
REGION Network 27: State 20 = Failed Ignition Attempt
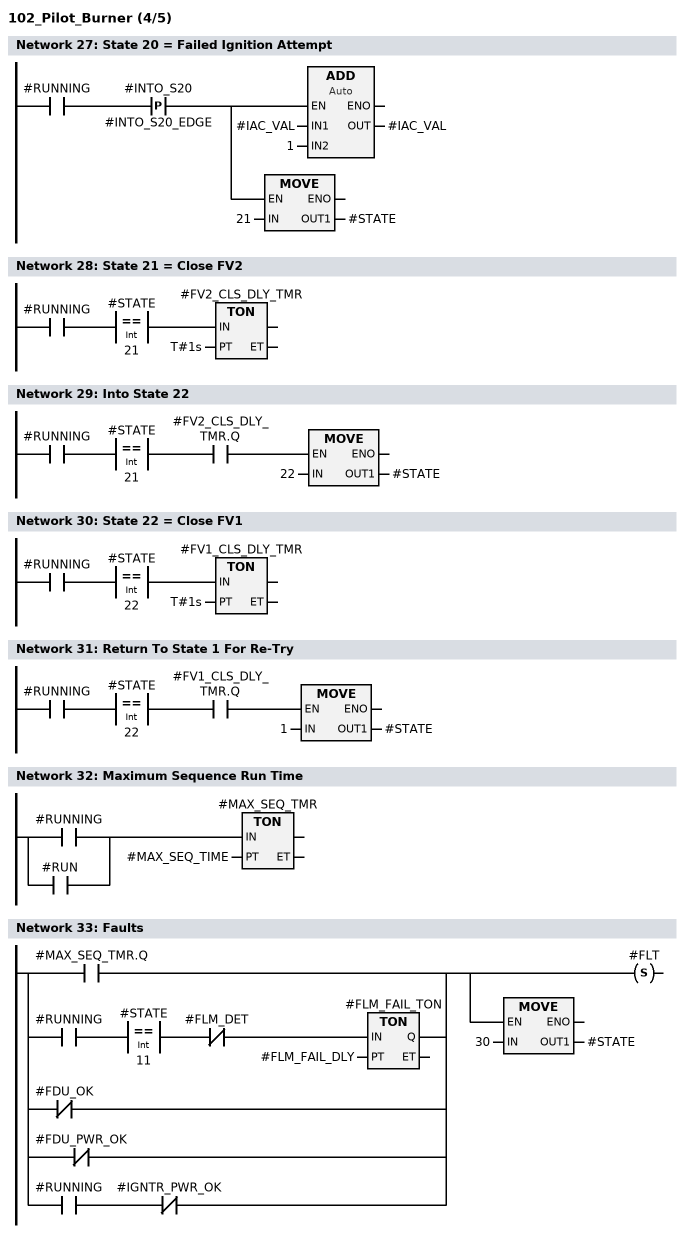
   RUNG wire#powerrail
      Contact( #RUNNING )
      P_Contact(operand := #INTO_S20, bit := #INTO_S20_EDGE)
      wire#w1
      Add(in1 := #IAC_VAL, in2 := 1, out => #IAC_VAL)
   END_RUNG
   RUNG wire#w1
      Move(in := 21, out1 => #STATE)
   END_RUNG
   // the same network as SCL:
   #_w1 := #RUNNING AND #INTO_S20 AND NOT #INTO_S20_EDGE;   // rising edge of #INTO_S20
   #INTO_S20_EDGE := #INTO_S20;
   IF #_w1 THEN
       #IAC_VAL := #IAC_VAL + 1;
       #STATE := 21;
   END_IF;
END_REGION

REGION Network 28: State 21 = Close FV2
   #FV2_CLS_DLY_TMR(IN := #RUNNING AND (#STATE = 21), PT := T#1s);   // TON
END_REGION

REGION Network 29: Into State 22
   RUNG wire#powerrail
      Contact( #RUNNING )
      { S7_Templates := "SrcType := Int" } EQ_Contact(in1 := #STATE, in2 := 21)
      Contact( #FV2_CLS_DLY_TMR.Q )
      Move(in := 22, out1 => #STATE)
   END_RUNG
   // the same network as SCL:
   IF #RUNNING AND (#STATE = 21) AND #FV2_CLS_DLY_TMR.Q THEN #STATE := 22; END_IF;
END_REGION

REGION Network 30: State 22 = Close FV1
   #FV1_CLS_DLY_TMR(IN := #RUNNING AND (#STATE = 22), PT := T#1s);   // TON
END_REGION

REGION Network 31: Return To State 1 For Re-Try
   RUNG wire#powerrail
      Contact( #RUNNING )
      { S7_Templates := "SrcType := Int" } EQ_Contact(in1 := #STATE, in2 := 22)
      Contact( #FV1_CLS_DLY_TMR.Q )
      Move(in := 1, out1 => #STATE)
   END_RUNG
   // the same network as SCL:
   IF #RUNNING AND (#STATE = 22) AND #FV1_CLS_DLY_TMR.Q THEN #STATE := 1; END_IF;
END_REGION

REGION Network 32: Maximum Sequence Run Time
   #MAX_SEQ_TMR(IN := #RUNNING OR #RUN, PT := #MAX_SEQ_TIME);   // TON
END_REGION

REGION Network 33: Faults
   #FLM_FAIL_TON(IN := #RUNNING AND (#STATE = 11) AND NOT #FLM_DET, PT := #FLM_FAIL_DLY);   // TON
   IF #MAX_SEQ_TMR.Q OR #FLM_FAIL_TON.Q OR NOT #FDU_OK OR NOT #FDU_PWR_OK OR (#RUNNING AND NOT #IGNTR_PWR_OK) THEN
       #FLT := TRUE;
       #STATE := 30;
   END_IF;
END_REGION

REGION Network 34: Reset Flag
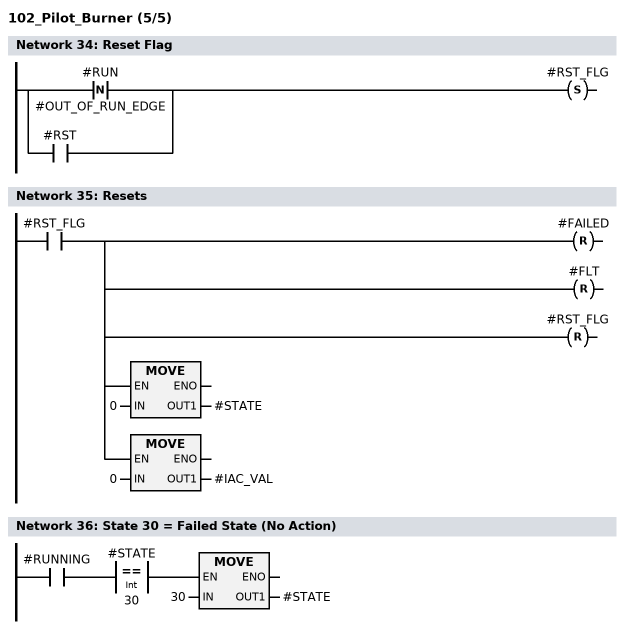
   RUNG wire#powerrail
      N_Contact(operand := #RUN, bit := #OUT_OF_RUN_EDGE)
      wire#w1
      S_Coil( #RST_FLG )
   END_RUNG
   RUNG wire#powerrail
      Contact( #RST )
   END_RUNG wire#w1
   // the same network as SCL:
   #_w1 := NOT #RUN AND #OUT_OF_RUN_EDGE;   // falling edge of #RUN
   #OUT_OF_RUN_EDGE := #RUN;
   IF #_w1 OR #RST THEN #RST_FLG := TRUE; END_IF;
END_REGION

REGION Network 35: Resets
   RUNG wire#powerrail
      Contact( #RST_FLG )
      wire#w1
      R_Coil( #FAILED )
   END_RUNG
   RUNG wire#w1
      R_Coil( #FLT )
   END_RUNG
   RUNG wire#w1
      R_Coil( #RST_FLG )
   END_RUNG
   RUNG wire#w1
      Move(in := 0, out1 => #STATE)
   END_RUNG
   RUNG wire#w1
      Move(in := 0, out1 => #IAC_VAL)
   END_RUNG
   // the same network as SCL:
   IF #RST_FLG THEN
       #FAILED := FALSE;
       #FLT := FALSE;
   END_IF;
   #_w1 := #RST_FLG;
   IF #_w1 THEN
       #RST_FLG := FALSE;
       #STATE := 0;
       #IAC_VAL := 0;
   END_IF;
END_REGION

REGION Network 36: State 30 = Failed State (No Action)
   RUNG wire#powerrail
      Contact( #RUNNING )
      { S7_Templates := "SrcType := Int" } EQ_Contact(in1 := #STATE, in2 := 30)
      Move(in := 30, out1 => #STATE)
   END_RUNG
   // the same network as SCL:
   IF #RUNNING AND (#STATE = 30) THEN #STATE := 30; END_IF;
END_REGION
END_FUNCTION_BLOCK

FUNCTION_BLOCK "103_Main_Burner"   // FB103, LAD
TITLE = Pilot Burner Control
{ S7_Optimized_Access := 'TRUE' }
AUTHOR : JRS
VERSION : 0.1
// For the control of the main burner ignition and burn
   VAR_INPUT
      RUN : Bool;   // Runs the block
      FLM_DET : Bool;   // Flame detected
      FLM_FAIL_DLY : Time;
      FV1_DLY : Time;   // Fuel valve 1 delay time
      FV2_3W_DLY : Time;   // 3 Way fuel valve 2 delay time
      FD_DLY : Time;   // Flame detection delay time
      FD_SCAN_TIME : Time;   // Flame detection scan time
      FD_VRFCTN_TIME : Time;   // Flame verification time
      MAX_SEQ_TIME : Time;   // Maximum sequence run time
      FDU_PWR_OK : Bool;   // Flame detection unit power ok
      FDU_OK : Bool;   // Flame detection health ok
      PrgdSTOP : Bool;
      RST : Bool;   // Reset bit
   END_VAR
   VAR_OUTPUT
      OPN_FV1 : Bool;   // Open fuel valve 1
      OPN_3W_FV2 : Bool;   // Open 3 way fuel valve 2
      DN_OK : Bool;   // Successful ignition
      FAILED : Bool;   // Ignition failed
      FLT : Bool;   // Fault bit
      Status : Int;
   END_VAR
   VAR_IN_OUT
      RUNNING : Bool;   // Sequence running
   END_VAR
   VAR
      INTO_RUN_EDGE : Bool;   // Edge detection
      OUT_OF_RUN_EDGE : Bool;   // Edge detection
      LOOK_NEG_EDGE : Bool;   // Stop looking edge
      INTO_S20 : Bool;   // Into step 20
      INTO_S20_EDGE : Bool;   // Into step 20 edge
      RST_FLG : Bool;   // Reset flag
      LOOKING : Bool;   // Looking for flame
      STATE : Int;   // State value for sequencing
      FD_SCN_TMR : TOF_TIME;   // Flame detection scan timer
      FV1_DLY_TMR : TON_TIME;   // Fuel valve 1 delay timer
      FV2_DLY_TMR : TON_TIME;   // Fuel valve 2 delay timer
      FD_DLY_TMR : TON_TIME;   // Flame detection delay timer
      FD_VRFCTN_TMR : TON_TIME;   // Flame verification timer
      MAX_SEQ_TMR : TON_TIME;   // Maximum sequence run timer
      FV1_CLS_DLY_TMR : TON_TIME;   // Fuel valve 1 close delay timer
      FV2_CLS_DLY_TMR : TON_TIME;   // Fuel valve 2 close delay timer
      IEC_Timer_0_Instance : TON_TIME;
      "Second beat" : TON_TIME;
   END_VAR
   VAR RETAIN
      "Seconds burn" : CTU_INT;
      "Minutes burn" : CTU_INT;
      "Hours burn" : CTU_INT;
      "Days burn" : CTU_INT;
      Aux : Struct
         Aux_1 : Bool;
         Aux_2 : Bool;
         Aux_3 : Bool;
         Aux_4 : Bool;
         AuxPulsReset : Bool;
      END_STRUCT;
   END_VAR
   VAR
      "Second Reset" : TON_TIME;
      "Not Run State" : TON_TIME;
      "Running TON" : TON_TIME;
      "Running State" : TON_TIME;
   END_VAR
   VAR_TEMP   // added for the SCL form of the ladder/FBD networks
      _w1 : Bool;
      _w2 : Bool;
      _w3 : Bool;
   END_VAR
BEGIN

REGION Network 1: Running
   // For running status detection
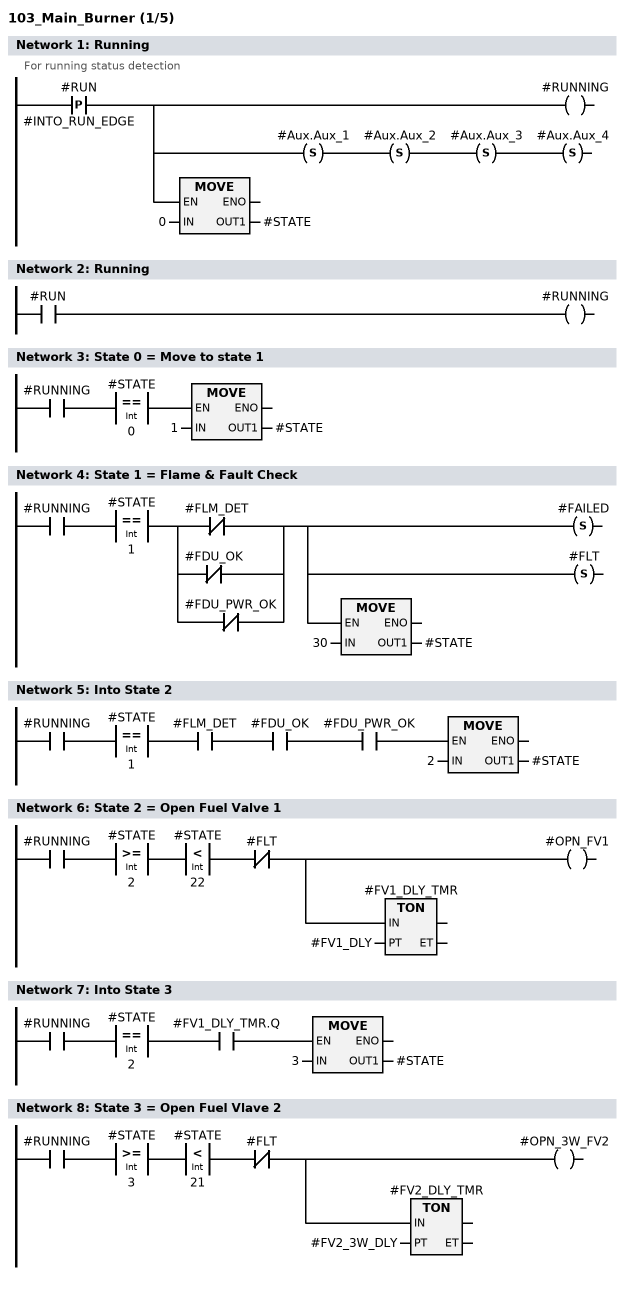
   RUNG wire#powerrail
      P_Contact(operand := #RUN, bit := #INTO_RUN_EDGE)
      wire#w1
      Coil( #RUNNING )
   END_RUNG
   RUNG wire#w1
      S_Coil( #Aux.Aux_1 )
      S_Coil( #Aux.Aux_2 )
      S_Coil( #Aux.Aux_3 )
      S_Coil( #Aux.Aux_4 )
   END_RUNG
   RUNG wire#w1
      Move(in := 0, out1 => #STATE)
   END_RUNG
   // the same network as SCL:
   #_w1 := #RUN AND NOT #INTO_RUN_EDGE;   // rising edge of #RUN
   #INTO_RUN_EDGE := #RUN;
   #RUNNING := #_w1;
   IF #_w1 THEN
       #Aux.Aux_1 := TRUE;
       #Aux.Aux_2 := TRUE;
       #Aux.Aux_3 := TRUE;
       #Aux.Aux_4 := TRUE;
       #STATE := 0;
   END_IF;
END_REGION

REGION Network 2: Running
   RUNG wire#powerrail
      Contact( #RUN )
      Coil( #RUNNING )
   END_RUNG
   // the same network as SCL:
   #RUNNING := #RUN;
END_REGION

REGION Network 3: State 0 = Move to state 1
   RUNG wire#powerrail
      Contact( #RUNNING )
      { S7_Templates := "SrcType := Int" } EQ_Contact(in1 := #STATE, in2 := 0)
      Move(in := 1, out1 => #STATE)
   END_RUNG
   // the same network as SCL:
   IF #RUNNING AND (#STATE = 0) THEN #STATE := 1; END_IF;
END_REGION

REGION Network 4: State 1 = Flame & Fault Check
   RUNG wire#powerrail
      Contact( #RUNNING )
      { S7_Templates := "SrcType := Int" } EQ_Contact(in1 := #STATE, in2 := 1)
      wire#w1
      I_Contact( #FLM_DET )
      wire#w2
      S_Coil( #FAILED )
   END_RUNG
   RUNG wire#w1
      I_Contact( #FDU_OK )
   END_RUNG wire#w2
   RUNG wire#w1
      I_Contact( #FDU_PWR_OK )
   END_RUNG wire#w2
   RUNG wire#w2
      S_Coil( #FLT )
   END_RUNG
   RUNG wire#w2
      Move(in := 30, out1 => #STATE)
   END_RUNG
   // the same network as SCL:
   IF #RUNNING AND (#STATE = 1) AND (NOT #FLM_DET OR NOT #FDU_OK OR NOT #FDU_PWR_OK) THEN
       #FAILED := TRUE;
       #FLT := TRUE;
       #STATE := 30;
   END_IF;
END_REGION

REGION Network 5: Into State 2
   RUNG wire#powerrail
      Contact( #RUNNING )
      { S7_Templates := "SrcType := Int" } EQ_Contact(in1 := #STATE, in2 := 1)
      Contact( #FLM_DET )
      Contact( #FDU_OK )
      Contact( #FDU_PWR_OK )
      Move(in := 2, out1 => #STATE)
   END_RUNG
   // the same network as SCL:
   IF #RUNNING AND (#STATE = 1) AND #FLM_DET AND #FDU_OK AND #FDU_PWR_OK THEN #STATE := 2; END_IF;
END_REGION

REGION Network 6: State 2 = Open Fuel Valve 1
   #OPN_FV1 := #RUNNING AND (#STATE >= 2) AND (#STATE < 22) AND NOT #FLT;
   #FV1_DLY_TMR(IN := #OPN_FV1, PT := #FV1_DLY);   // TON
END_REGION

REGION Network 7: Into State 3
   RUNG wire#powerrail
      Contact( #RUNNING )
      { S7_Templates := "SrcType := Int" } EQ_Contact(in1 := #STATE, in2 := 2)
      Contact( #FV1_DLY_TMR.Q )
      Move(in := 3, out1 => #STATE)
   END_RUNG
   // the same network as SCL:
   IF #RUNNING AND (#STATE = 2) AND #FV1_DLY_TMR.Q THEN #STATE := 3; END_IF;
END_REGION

REGION Network 8: State 3 = Open Fuel Vlave 2
   #OPN_3W_FV2 := #RUNNING AND (#STATE >= 3) AND (#STATE < 21) AND NOT #FLT;
   #FV2_DLY_TMR(IN := #OPN_3W_FV2, PT := #FV2_3W_DLY);   // TON
END_REGION

REGION Network 9: Into State 4
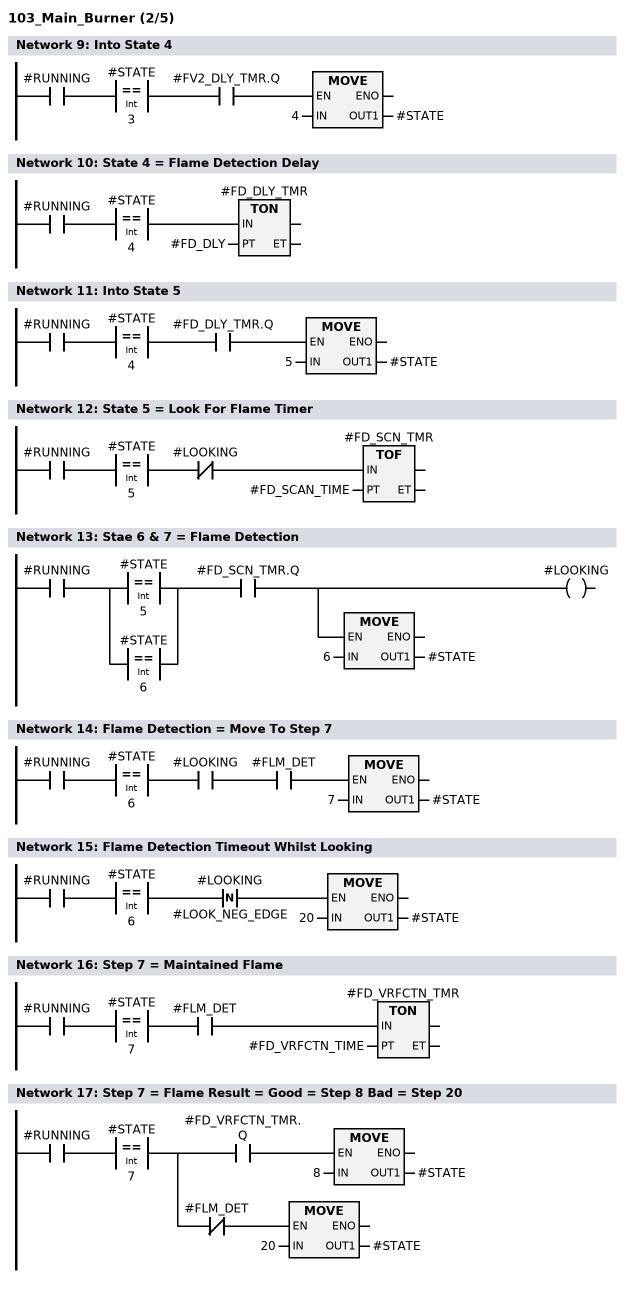
   RUNG wire#powerrail
      Contact( #RUNNING )
      { S7_Templates := "SrcType := Int" } EQ_Contact(in1 := #STATE, in2 := 3)
      Contact( #FV2_DLY_TMR.Q )
      Move(in := 4, out1 => #STATE)
   END_RUNG
   // the same network as SCL:
   IF #RUNNING AND (#STATE = 3) AND #FV2_DLY_TMR.Q THEN #STATE := 4; END_IF;
END_REGION

REGION Network 10: State 4 = Flame Detection Delay
   #FD_DLY_TMR(IN := #RUNNING AND (#STATE = 4), PT := #FD_DLY);   // TON
END_REGION

REGION Network 11: Into State 5
   RUNG wire#powerrail
      Contact( #RUNNING )
      { S7_Templates := "SrcType := Int" } EQ_Contact(in1 := #STATE, in2 := 4)
      Contact( #FD_DLY_TMR.Q )
      Move(in := 5, out1 => #STATE)
   END_RUNG
   // the same network as SCL:
   IF #RUNNING AND (#STATE = 4) AND #FD_DLY_TMR.Q THEN #STATE := 5; END_IF;
END_REGION

REGION Network 12: State 5 = Look For Flame Timer
   #FD_SCN_TMR(IN := #RUNNING AND (#STATE = 5) AND NOT #LOOKING, PT := #FD_SCAN_TIME);   // TOF
END_REGION

REGION Network 13: Stae 6 & 7 = Flame Detection
   RUNG wire#powerrail
      Contact( #RUNNING )
      wire#w1
      { S7_Templates := "SrcType := Int" } EQ_Contact(in1 := #STATE, in2 := 5)
      wire#w2
      Contact( #FD_SCN_TMR.Q )
      wire#w3
      Coil( #LOOKING )
   END_RUNG
   RUNG wire#w1
      { S7_Templates := "SrcType := Int" } EQ_Contact(in1 := #STATE, in2 := 6)
   END_RUNG wire#w2
   RUNG wire#w3
      Move(in := 6, out1 => #STATE)
   END_RUNG
   // the same network as SCL:
   #LOOKING := #RUNNING AND ((#STATE = 5) OR (#STATE = 6)) AND #FD_SCN_TMR.Q;
   IF #LOOKING THEN #STATE := 6; END_IF;
END_REGION

REGION Network 14: Flame Detection = Move To Step 7
   RUNG wire#powerrail
      Contact( #RUNNING )
      { S7_Templates := "SrcType := Int" } EQ_Contact(in1 := #STATE, in2 := 6)
      Contact( #LOOKING )
      Contact( #FLM_DET )
      Move(in := 7, out1 => #STATE)
   END_RUNG
   // the same network as SCL:
   IF #RUNNING AND (#STATE = 6) AND #LOOKING AND #FLM_DET THEN #STATE := 7; END_IF;
END_REGION

REGION Network 15: Flame Detection Timeout Whilst Looking
   RUNG wire#powerrail
      Contact( #RUNNING )
      { S7_Templates := "SrcType := Int" } EQ_Contact(in1 := #STATE, in2 := 6)
      N_Contact(operand := #LOOKING, bit := #LOOK_NEG_EDGE)
      Move(in := 20, out1 => #STATE)
   END_RUNG
   // the same network as SCL:
   #_w1 := #RUNNING AND (#STATE = 6) AND NOT #LOOKING AND #LOOK_NEG_EDGE;   // falling edge of #LOOKING
   #LOOK_NEG_EDGE := #LOOKING;
   IF #_w1 THEN #STATE := 20; END_IF;
END_REGION

REGION Network 16: Step 7 = Maintained Flame
   #FD_VRFCTN_TMR(IN := #RUNNING AND (#STATE = 7) AND #FLM_DET, PT := #FD_VRFCTN_TIME);   // TON
END_REGION

REGION Network 17: Step 7 = Flame Result = Good = Step 8 Bad = Step 20
   RUNG wire#powerrail
      Contact( #RUNNING )
      { S7_Templates := "SrcType := Int" } EQ_Contact(in1 := #STATE, in2 := 7)
      wire#w1
      Contact( #FD_VRFCTN_TMR.Q )
      Move(in := 8, out1 => #STATE)
   END_RUNG
   RUNG wire#w1
      I_Contact( #FLM_DET )
      Move(in := 20, out1 => #STATE)
   END_RUNG
   // the same network as SCL:
   #_w1 := #RUNNING AND (#STATE = 7);
   IF #_w1 AND #FD_VRFCTN_TMR.Q THEN #STATE := 8; END_IF;
   IF #_w1 AND NOT #FLM_DET THEN #STATE := 20; END_IF;
END_REGION

REGION Network 18: State 8 = Check Flame Still Detected
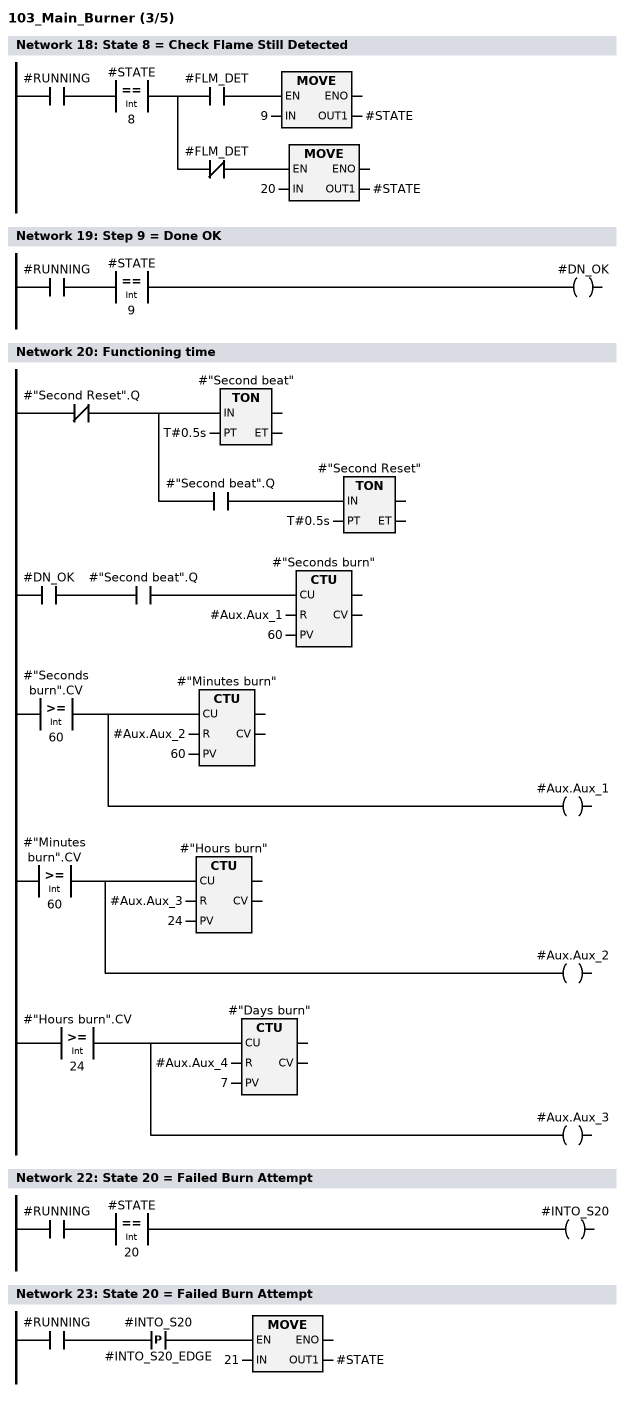
   RUNG wire#powerrail
      Contact( #RUNNING )
      { S7_Templates := "SrcType := Int" } EQ_Contact(in1 := #STATE, in2 := 8)
      wire#w1
      Contact( #FLM_DET )
      Move(in := 9, out1 => #STATE)
   END_RUNG
   RUNG wire#w1
      I_Contact( #FLM_DET )
      Move(in := 20, out1 => #STATE)
   END_RUNG
   // the same network as SCL:
   #_w1 := #RUNNING AND (#STATE = 8);
   IF #_w1 AND #FLM_DET THEN #STATE := 9; END_IF;
   IF #_w1 AND NOT #FLM_DET THEN #STATE := 20; END_IF;
END_REGION

REGION Network 19: Step 9 = Done OK
   RUNG wire#powerrail
      Contact( #RUNNING )
      { S7_Templates := "SrcType := Int" } EQ_Contact(in1 := #STATE, in2 := 9)
      Coil( #DN_OK )
   END_RUNG
   // the same network as SCL:
   #DN_OK := #RUNNING AND (#STATE = 9);
END_REGION

REGION Network 20: Functioning time
   #"Second beat"(IN := NOT #"Second Reset".Q, PT := T#0.5s);   // TON
   #"Second Reset"(IN := NOT #"Second Reset".Q AND #"Second beat".Q, PT := T#0.5s);   // TON
   #"Seconds burn"(CU := #DN_OK AND #"Second beat".Q, R := #Aux.Aux_1, PV := 60);   // CTU
   #_w1 := #"Seconds burn".CV >= 60;
   #"Minutes burn"(CU := #_w1, R := #Aux.Aux_2, PV := 60);   // CTU
   #Aux.Aux_1 := #_w1;
   #_w2 := #"Minutes burn".CV >= 60;
   #"Hours burn"(CU := #_w2, R := #Aux.Aux_3, PV := 24);   // CTU
   #Aux.Aux_2 := #_w2;
   #_w3 := #"Hours burn".CV >= 24;
   #"Days burn"(CU := #_w3, R := #Aux.Aux_4, PV := 7);   // CTU
   #Aux.Aux_3 := #_w3;
END_REGION

REGION Network 22: State 20 = Failed Burn Attempt
   RUNG wire#powerrail
      Contact( #RUNNING )
      { S7_Templates := "SrcType := Int" } EQ_Contact(in1 := #STATE, in2 := 20)
      Coil( #INTO_S20 )
   END_RUNG
   // the same network as SCL:
   #INTO_S20 := #RUNNING AND (#STATE = 20);
END_REGION

REGION Network 23: State 20 = Failed Burn Attempt
   RUNG wire#powerrail
      Contact( #RUNNING )
      P_Contact(operand := #INTO_S20, bit := #INTO_S20_EDGE)
      Move(in := 21, out1 => #STATE)
   END_RUNG
   // the same network as SCL:
   #_w1 := #RUNNING AND #INTO_S20 AND NOT #INTO_S20_EDGE;   // rising edge of #INTO_S20
   #INTO_S20_EDGE := #INTO_S20;
   IF #_w1 THEN #STATE := 21; END_IF;
END_REGION

REGION Network 24: State 21 = Close FV2
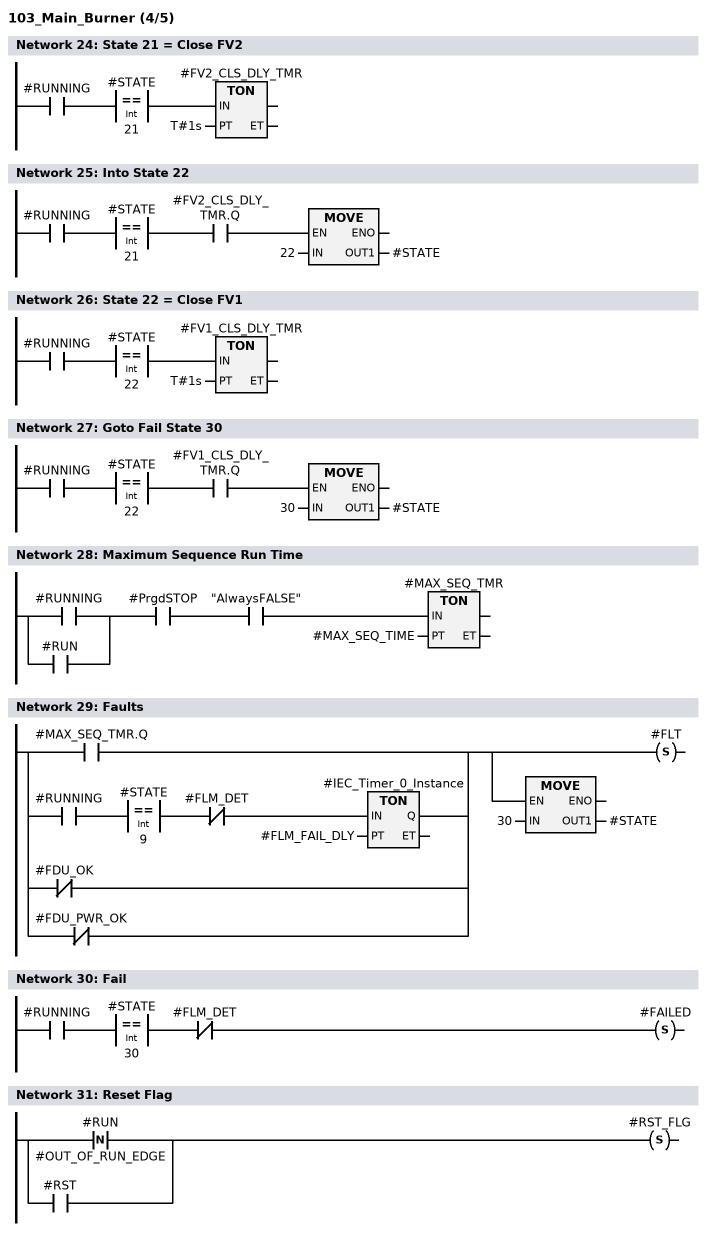
   #FV2_CLS_DLY_TMR(IN := #RUNNING AND (#STATE = 21), PT := T#1s);   // TON
END_REGION

REGION Network 25: Into State 22
   RUNG wire#powerrail
      Contact( #RUNNING )
      { S7_Templates := "SrcType := Int" } EQ_Contact(in1 := #STATE, in2 := 21)
      Contact( #FV2_CLS_DLY_TMR.Q )
      Move(in := 22, out1 => #STATE)
   END_RUNG
   // the same network as SCL:
   IF #RUNNING AND (#STATE = 21) AND #FV2_CLS_DLY_TMR.Q THEN #STATE := 22; END_IF;
END_REGION

REGION Network 26: State 22 = Close FV1
   #FV1_CLS_DLY_TMR(IN := #RUNNING AND (#STATE = 22), PT := T#1s);   // TON
END_REGION

REGION Network 27: Goto Fail State 30
   RUNG wire#powerrail
      Contact( #RUNNING )
      { S7_Templates := "SrcType := Int" } EQ_Contact(in1 := #STATE, in2 := 22)
      Contact( #FV1_CLS_DLY_TMR.Q )
      Move(in := 30, out1 => #STATE)
   END_RUNG
   // the same network as SCL:
   IF #RUNNING AND (#STATE = 22) AND #FV1_CLS_DLY_TMR.Q THEN #STATE := 30; END_IF;
END_REGION

REGION Network 28: Maximum Sequence Run Time
   #MAX_SEQ_TMR(IN := (#RUNNING OR #RUN) AND #PrgdSTOP AND "AlwaysFALSE", PT := #MAX_SEQ_TIME);   // TON
END_REGION

REGION Network 29: Faults
   #IEC_Timer_0_Instance(IN := #RUNNING AND (#STATE = 9) AND NOT #FLM_DET, PT := #FLM_FAIL_DLY);   // TON
   IF #MAX_SEQ_TMR.Q OR #IEC_Timer_0_Instance.Q OR NOT #FDU_OK OR NOT #FDU_PWR_OK THEN
       #FLT := TRUE;
       #STATE := 30;
   END_IF;
END_REGION

REGION Network 30: Fail
   RUNG wire#powerrail
      Contact( #RUNNING )
      { S7_Templates := "SrcType := Int" } EQ_Contact(in1 := #STATE, in2 := 30)
      I_Contact( #FLM_DET )
      S_Coil( #FAILED )
   END_RUNG
   // the same network as SCL:
   IF #RUNNING AND (#STATE = 30) AND NOT #FLM_DET THEN #FAILED := TRUE; END_IF;
END_REGION

REGION Network 31: Reset Flag
   RUNG wire#powerrail
      N_Contact(operand := #RUN, bit := #OUT_OF_RUN_EDGE)
      wire#w1
      S_Coil( #RST_FLG )
   END_RUNG
   RUNG wire#powerrail
      Contact( #RST )
   END_RUNG wire#w1
   // the same network as SCL:
   #_w1 := NOT #RUN AND #OUT_OF_RUN_EDGE;   // falling edge of #RUN
   #OUT_OF_RUN_EDGE := #RUN;
   IF #_w1 OR #RST THEN #RST_FLG := TRUE; END_IF;
END_REGION

REGION Network 32: Resets
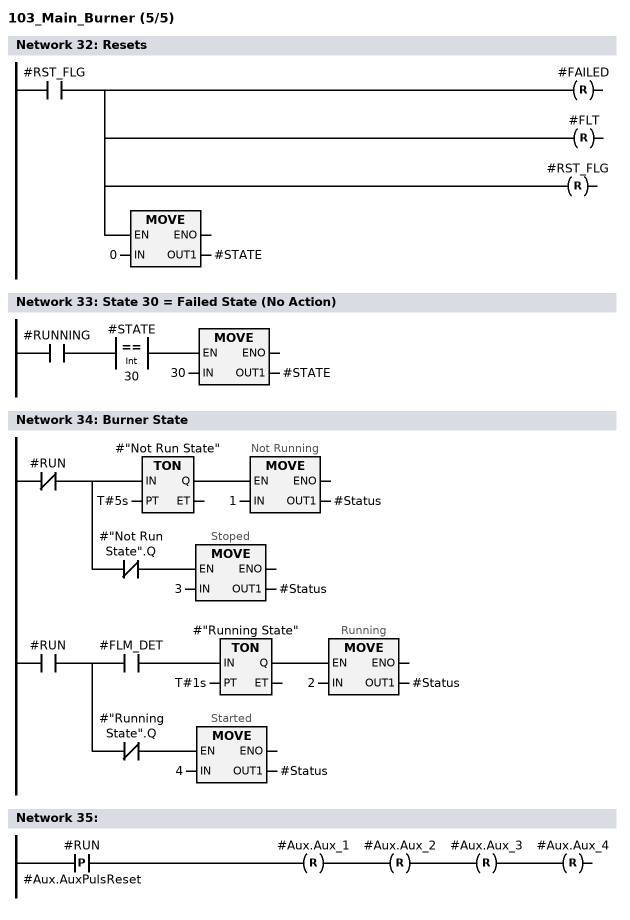
   RUNG wire#powerrail
      Contact( #RST_FLG )
      wire#w1
      R_Coil( #FAILED )
   END_RUNG
   RUNG wire#w1
      R_Coil( #FLT )
   END_RUNG
   RUNG wire#w1
      R_Coil( #RST_FLG )
   END_RUNG
   RUNG wire#w1
      Move(in := 0, out1 => #STATE)
   END_RUNG
   // the same network as SCL:
   IF #RST_FLG THEN
       #FAILED := FALSE;
       #FLT := FALSE;
   END_IF;
   #_w1 := #RST_FLG;
   IF #_w1 THEN
       #RST_FLG := FALSE;
       #STATE := 0;
   END_IF;
END_REGION

REGION Network 33: State 30 = Failed State (No Action)
   RUNG wire#powerrail
      Contact( #RUNNING )
      { S7_Templates := "SrcType := Int" } EQ_Contact(in1 := #STATE, in2 := 30)
      Move(in := 30, out1 => #STATE)
   END_RUNG
   // the same network as SCL:
   IF #RUNNING AND (#STATE = 30) THEN #STATE := 30; END_IF;
END_REGION

REGION Network 34: Burner State
   #"Not Run State"(IN := NOT #RUN, PT := T#5s);   // TON
   IF #"Not Run State".Q THEN
       #Status := 1;   // Not Running
   END_IF;
   IF NOT #RUN AND NOT #"Not Run State".Q THEN
       #Status := 3;   // Stoped
   END_IF;
   #"Running State"(IN := #RUN AND #FLM_DET, PT := T#1s);   // TON
   IF #"Running State".Q THEN
       #Status := 2;   // Running
   END_IF;
   IF #RUN AND NOT #"Running State".Q THEN
       #Status := 4;   // Started
   END_IF;
END_REGION

REGION Network 35
   RUNG wire#powerrail
      P_Contact(operand := #RUN, bit := #Aux.AuxPulsReset)
      R_Coil( #Aux.Aux_1 )
      R_Coil( #Aux.Aux_2 )
      R_Coil( #Aux.Aux_3 )
      R_Coil( #Aux.Aux_4 )
   END_RUNG
   // the same network as SCL:
   #_w1 := #RUN AND NOT #Aux.AuxPulsReset;   // rising edge of #RUN
   #Aux.AuxPulsReset := #RUN;
   IF #_w1 THEN
       #Aux.Aux_1 := FALSE;
       #Aux.Aux_2 := FALSE;
       #Aux.Aux_3 := FALSE;
       #Aux.Aux_4 := FALSE;
   END_IF;
END_REGION
END_FUNCTION_BLOCK

FUNCTION_BLOCK "104_Pilot_Purge"   // FB104, LAD
TITLE = Pilot Burner Purge
{ S7_Optimized_Access := 'TRUE' }
AUTHOR : JRS
VERSION : 0.1
// For the control of the pilot burner purge sequence
   VAR_INPUT
      RUN : Bool;   // Runs the block
      AV_Q : Bool;   // Air valve output state
      FV1_Q : Bool;   // Fuel valve 1 output state
      FV2_3W_Q : Bool;   // 3 Way fuel valve 2 output state
      FV1_CLS_DLY : Time;   // Fuel valve 1 delay time
      FV2_3W_CLS_DLY : Time;   // 3 Way fuel valve 2 delay time
      FV2_3W_OPN_DLY : Time;   // 3 Way fuel valve 2 delay time
      AV_CLS_DLY : Time;   // Air valve delay time
      MAX_SEQ_TIME : Time;   // Maximum sequence run time
      RST : Bool;   // Reset bit
   END_VAR
   VAR_OUTPUT
      PRG_ACTV : Bool;   // Purge active
      OPN_AV : Bool;   // Open air valve
      OPN_FV1 : Bool;   // Open fuel valve 1
      OPN_3W_FV2 : Bool;   // Open 3 way fuel valve 2
      DN_OK : Bool;   // Successful ignition
      FLT : Bool;   // Fault bit
   END_VAR
   VAR_IN_OUT
      RUNNING : Bool;   // Sequence running
   END_VAR
   VAR
      INTO_RUN_EDGE : Bool;   // Edge detection
      OUT_OF_RUN_EDGE : Bool;   // Edge detection
      RST_FLG : Bool;   // Reset flag
      ACTIVE : Bool;   // Active flag
      STATE : Int;   // State value for sequencing
      FV1_DLY_TMR : TON_TIME;   // Fuel valve 1 delay timer
      FV2_DLY_TMR : TON_TIME;   // Fuel valve 2 delay timer
      AV_DLY_TMR : TON_TIME;   // Air valve delay timer
      MAX_SEQ_TMR : TON_TIME;   // Maximum sequence run timer
      FV2_OPN_DLY_TMR : TON_TIME;   // Fuel valve 2 open delay timer
   END_VAR
   VAR_TEMP   // added for the SCL form of the ladder/FBD networks
      _w1 : Bool;
   END_VAR
BEGIN

REGION Network 1: Running
   // For running status detection
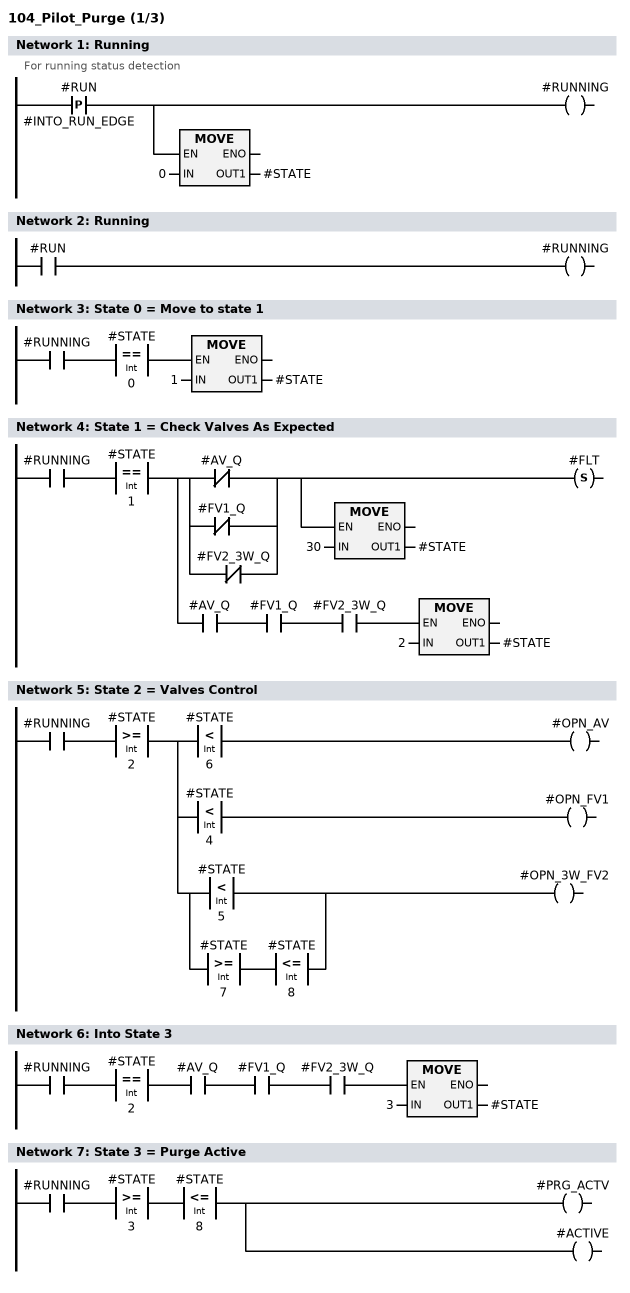
   RUNG wire#powerrail
      P_Contact(operand := #RUN, bit := #INTO_RUN_EDGE)
      wire#w1
      Coil( #RUNNING )
   END_RUNG
   RUNG wire#w1
      Move(in := 0, out1 => #STATE)
   END_RUNG
   // the same network as SCL:
   #_w1 := #RUN AND NOT #INTO_RUN_EDGE;   // rising edge of #RUN
   #INTO_RUN_EDGE := #RUN;
   #RUNNING := #_w1;
   IF #_w1 THEN #STATE := 0; END_IF;
END_REGION

REGION Network 2: Running
   RUNG wire#powerrail
      Contact( #RUN )
      Coil( #RUNNING )
   END_RUNG
   // the same network as SCL:
   #RUNNING := #RUN;
END_REGION

REGION Network 3: State 0 = Move to state 1
   RUNG wire#powerrail
      Contact( #RUNNING )
      { S7_Templates := "SrcType := Int" } EQ_Contact(in1 := #STATE, in2 := 0)
      Move(in := 1, out1 => #STATE)
   END_RUNG
   // the same network as SCL:
   IF #RUNNING AND (#STATE = 0) THEN #STATE := 1; END_IF;
END_REGION

REGION Network 4: State 1 = Check Valves As Expected
   RUNG wire#powerrail
      Contact( #RUNNING )
      { S7_Templates := "SrcType := Int" } EQ_Contact(in1 := #STATE, in2 := 1)
      wire#w1
      I_Contact( #AV_Q )
      wire#w2
      S_Coil( #FLT )
   END_RUNG
   RUNG wire#w1
      I_Contact( #FV1_Q )
   END_RUNG wire#w2
   RUNG wire#w1
      I_Contact( #FV2_3W_Q )
   END_RUNG wire#w2
   RUNG wire#w2
      Move(in := 30, out1 => #STATE)
   END_RUNG
   RUNG wire#w1
      Contact( #AV_Q )
      Contact( #FV1_Q )
      Contact( #FV2_3W_Q )
      Move(in := 2, out1 => #STATE)
   END_RUNG
   // the same network as SCL:
   #_w1 := #RUNNING AND (#STATE = 1);
   IF #_w1 AND (NOT #AV_Q OR NOT #FV1_Q OR NOT #FV2_3W_Q) THEN
       #FLT := TRUE;
       #STATE := 30;
   END_IF;
   IF #_w1 AND #AV_Q AND #FV1_Q AND #FV2_3W_Q THEN #STATE := 2; END_IF;
END_REGION
